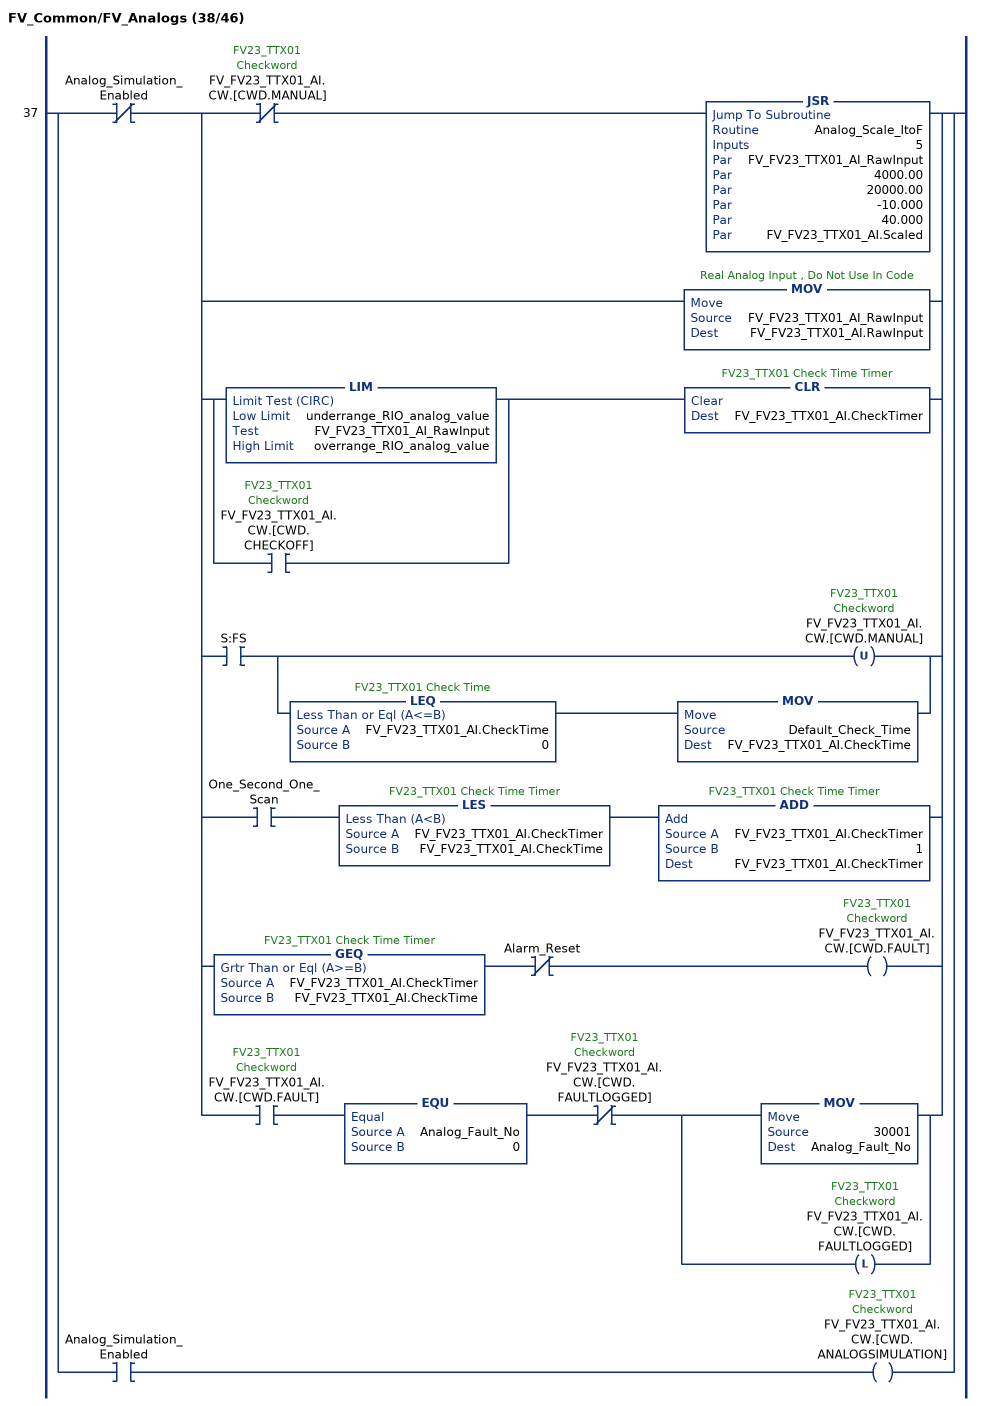
   37: [XIO(Analog_Simulation_Enabled) [XIO(FV_FV23_TTX01_AI.CW.[CWD.MANUAL]) JSR(Analog_Scale_ItoF,5,FV_FV23_TTX01_AI_RawInput,4000.00,20000.00,-10.000,40.000,FV_FV23_TTX01_AI.Scaled) ,MOV(FV_FV23_TTX01_AI_RawInput,FV_FV23_TTX01_AI.RawInput) ,[LIM(underrange_RIO_analog_value,FV_FV23_TTX01_AI_RawInput,overrange_RIO_analog_value) ,XIC(FV_FV23_TTX01_AI.CW.[CWD.CHECKOFF]) ] CLR(FV_FV23_TTX01_AI.CheckTimer) ,XIC(S:FS) [OTU(FV_FV23_TTX01_AI.CW.[CWD.MANUAL]) ,LEQ(FV_FV23_TTX01_AI.CheckTime,0) MOV(Default_Check_Time,FV_FV23_TTX01_AI.CheckTime) ] ,XIC(One_Second_One_Scan) LES(FV_FV23_TTX01_AI.CheckTimer,FV_FV23_TTX01_AI.CheckTime) ADD(FV_FV23_TTX01_AI.CheckTimer,1,FV_FV23_TTX01_AI.CheckTimer) ,GEQ(FV_FV23_TTX01_AI.CheckTimer,FV_FV23_TTX01_AI.CheckTime) XIO(Alarm_Reset) OTE(FV_FV23_TTX01_AI.CW.[CWD.FAULT]) ,XIC(FV_FV23_TTX01_AI.CW.[CWD.FAULT]) EQU(Analog_Fault_No,0) XIO(FV_FV23_TTX01_AI.CW.[CWD.FAULTLOGGED]) [MOV(30001,Analog_Fault_No) ,OTL(FV_FV23_TTX01_AI.CW.[CWD.FAULTLOGGED]) ] ] ,XIC(Analog_Simulation_Enabled) OTE(FV_FV23_TTX01_AI.CW.[CWD.ANALOGSIMULATION]) ];
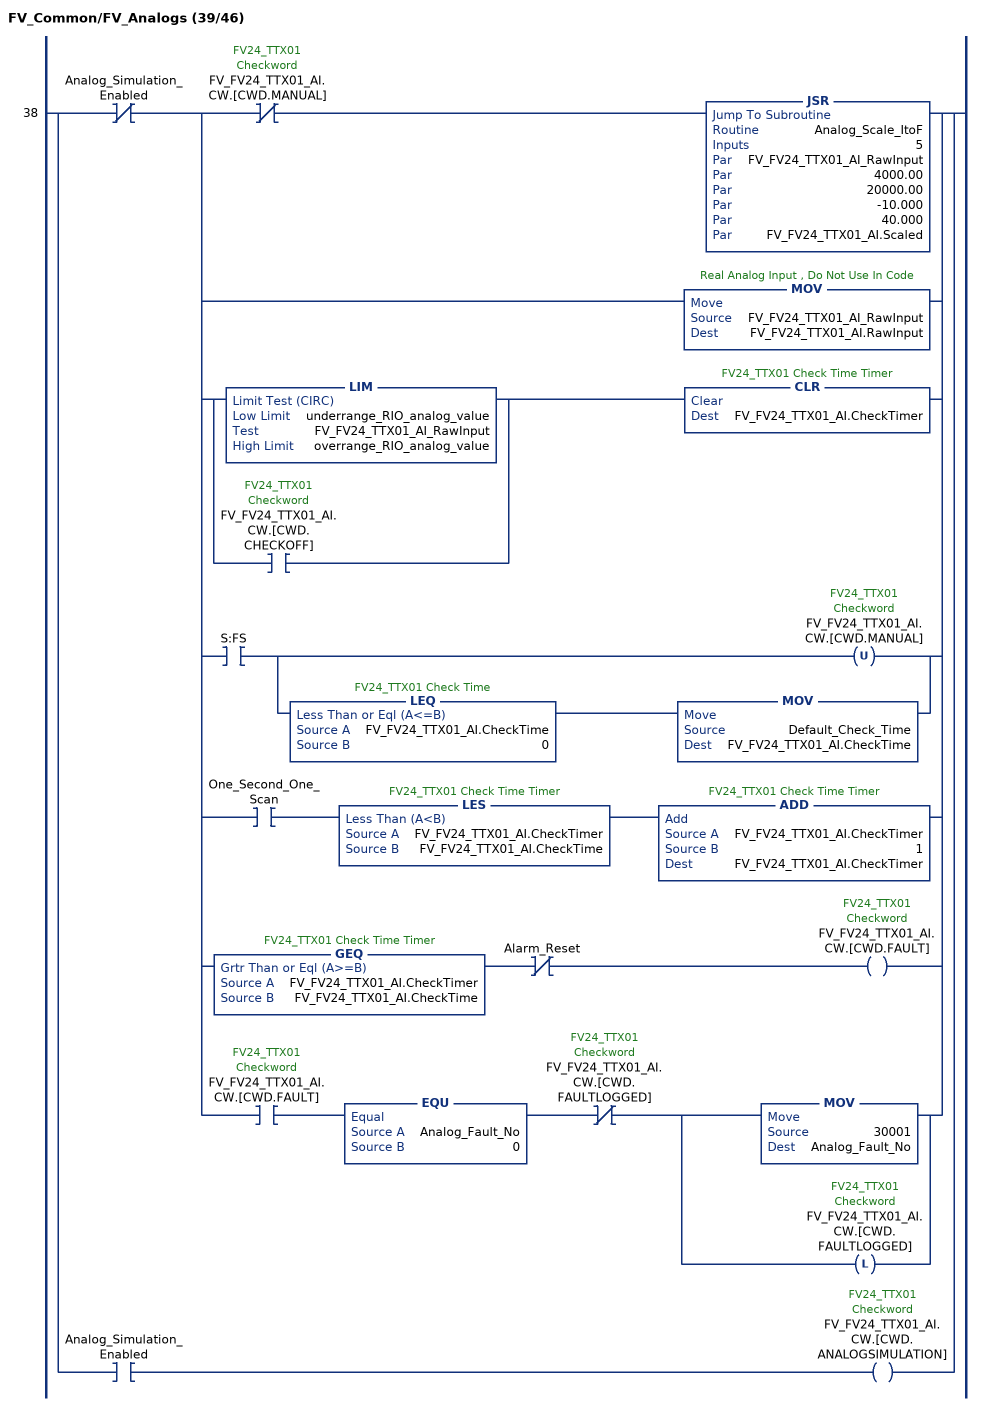
   38: [XIO(Analog_Simulation_Enabled) [XIO(FV_FV24_TTX01_AI.CW.[CWD.MANUAL]) JSR(Analog_Scale_ItoF,5,FV_FV24_TTX01_AI_RawInput,4000.00,20000.00,-10.000,40.000,FV_FV24_TTX01_AI.Scaled) ,MOV(FV_FV24_TTX01_AI_RawInput,FV_FV24_TTX01_AI.RawInput) ,[LIM(underrange_RIO_analog_value,FV_FV24_TTX01_AI_RawInput,overrange_RIO_analog_value) ,XIC(FV_FV24_TTX01_AI.CW.[CWD.CHECKOFF]) ] CLR(FV_FV24_TTX01_AI.CheckTimer) ,XIC(S:FS) [OTU(FV_FV24_TTX01_AI.CW.[CWD.MANUAL]) ,LEQ(FV_FV24_TTX01_AI.CheckTime,0) MOV(Default_Check_Time,FV_FV24_TTX01_AI.CheckTime) ] ,XIC(One_Second_One_Scan) LES(FV_FV24_TTX01_AI.CheckTimer,FV_FV24_TTX01_AI.CheckTime) ADD(FV_FV24_TTX01_AI.CheckTimer,1,FV_FV24_TTX01_AI.CheckTimer) ,GEQ(FV_FV24_TTX01_AI.CheckTimer,FV_FV24_TTX01_AI.CheckTime) XIO(Alarm_Reset) OTE(FV_FV24_TTX01_AI.CW.[CWD.FAULT]) ,XIC(FV_FV24_TTX01_AI.CW.[CWD.FAULT]) EQU(Analog_Fault_No,0) XIO(FV_FV24_TTX01_AI.CW.[CWD.FAULTLOGGED]) [MOV(30001,Analog_Fault_No) ,OTL(FV_FV24_TTX01_AI.CW.[CWD.FAULTLOGGED]) ] ] ,XIC(Analog_Simulation_Enabled) OTE(FV_FV24_TTX01_AI.CW.[CWD.ANALOGSIMULATION]) ];
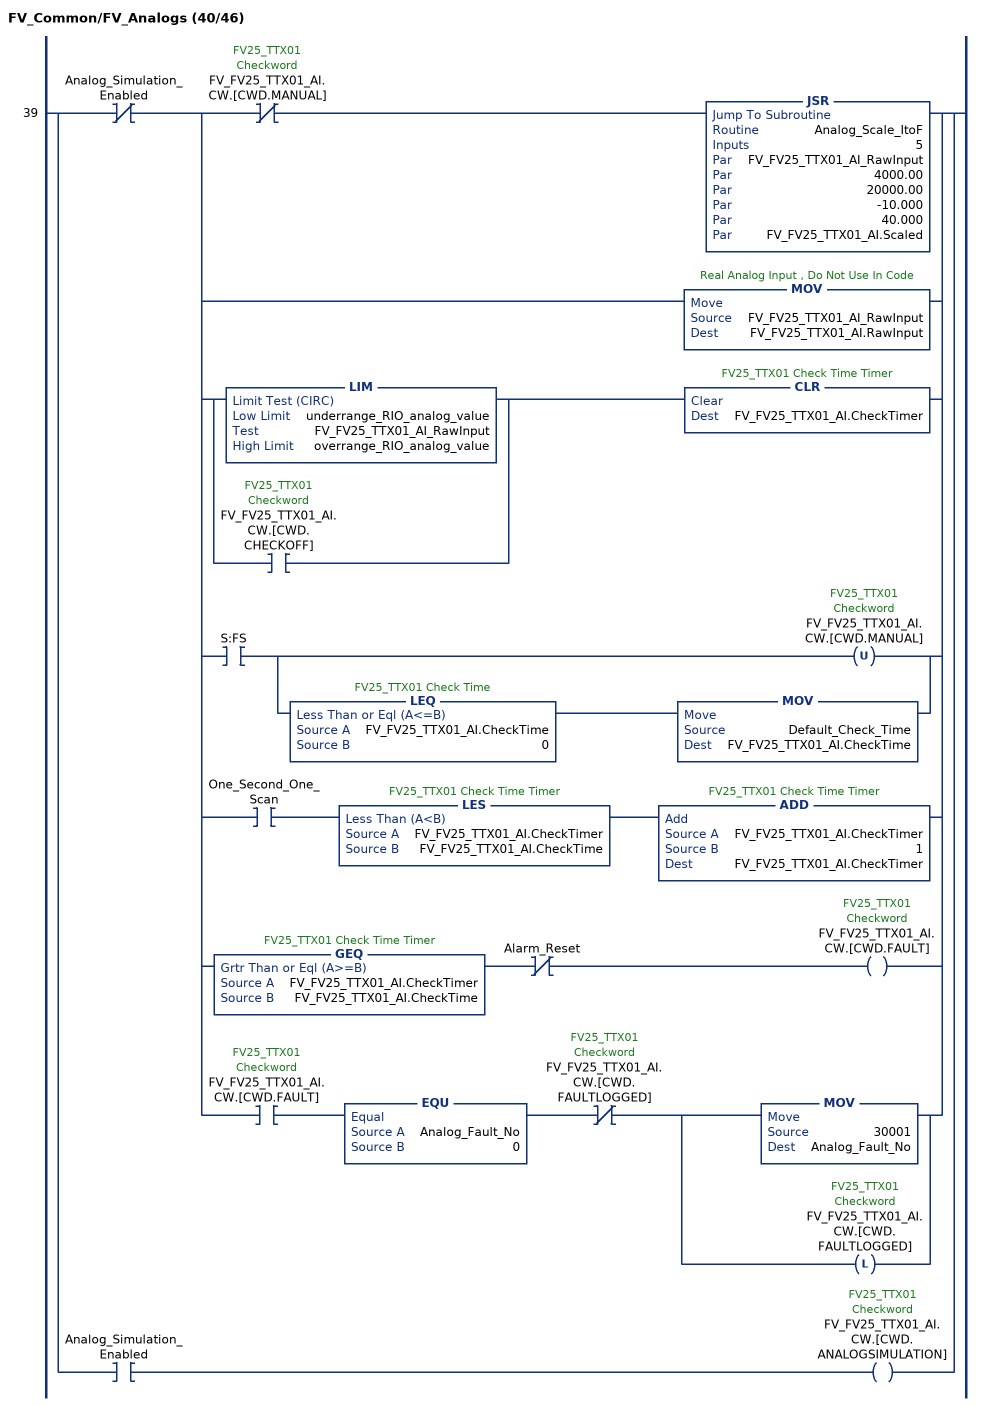
   39: [XIO(Analog_Simulation_Enabled) [XIO(FV_FV25_TTX01_AI.CW.[CWD.MANUAL]) JSR(Analog_Scale_ItoF,5,FV_FV25_TTX01_AI_RawInput,4000.00,20000.00,-10.000,40.000,FV_FV25_TTX01_AI.Scaled) ,MOV(FV_FV25_TTX01_AI_RawInput,FV_FV25_TTX01_AI.RawInput) ,[LIM(underrange_RIO_analog_value,FV_FV25_TTX01_AI_RawInput,overrange_RIO_analog_value) ,XIC(FV_FV25_TTX01_AI.CW.[CWD.CHECKOFF]) ] CLR(FV_FV25_TTX01_AI.CheckTimer) ,XIC(S:FS) [OTU(FV_FV25_TTX01_AI.CW.[CWD.MANUAL]) ,LEQ(FV_FV25_TTX01_AI.CheckTime,0) MOV(Default_Check_Time,FV_FV25_TTX01_AI.CheckTime) ] ,XIC(One_Second_One_Scan) LES(FV_FV25_TTX01_AI.CheckTimer,FV_FV25_TTX01_AI.CheckTime) ADD(FV_FV25_TTX01_AI.CheckTimer,1,FV_FV25_TTX01_AI.CheckTimer) ,GEQ(FV_FV25_TTX01_AI.CheckTimer,FV_FV25_TTX01_AI.CheckTime) XIO(Alarm_Reset) OTE(FV_FV25_TTX01_AI.CW.[CWD.FAULT]) ,XIC(FV_FV25_TTX01_AI.CW.[CWD.FAULT]) EQU(Analog_Fault_No,0) XIO(FV_FV25_TTX01_AI.CW.[CWD.FAULTLOGGED]) [MOV(30001,Analog_Fault_No) ,OTL(FV_FV25_TTX01_AI.CW.[CWD.FAULTLOGGED]) ] ] ,XIC(Analog_Simulation_Enabled) OTE(FV_FV25_TTX01_AI.CW.[CWD.ANALOGSIMULATION]) ];
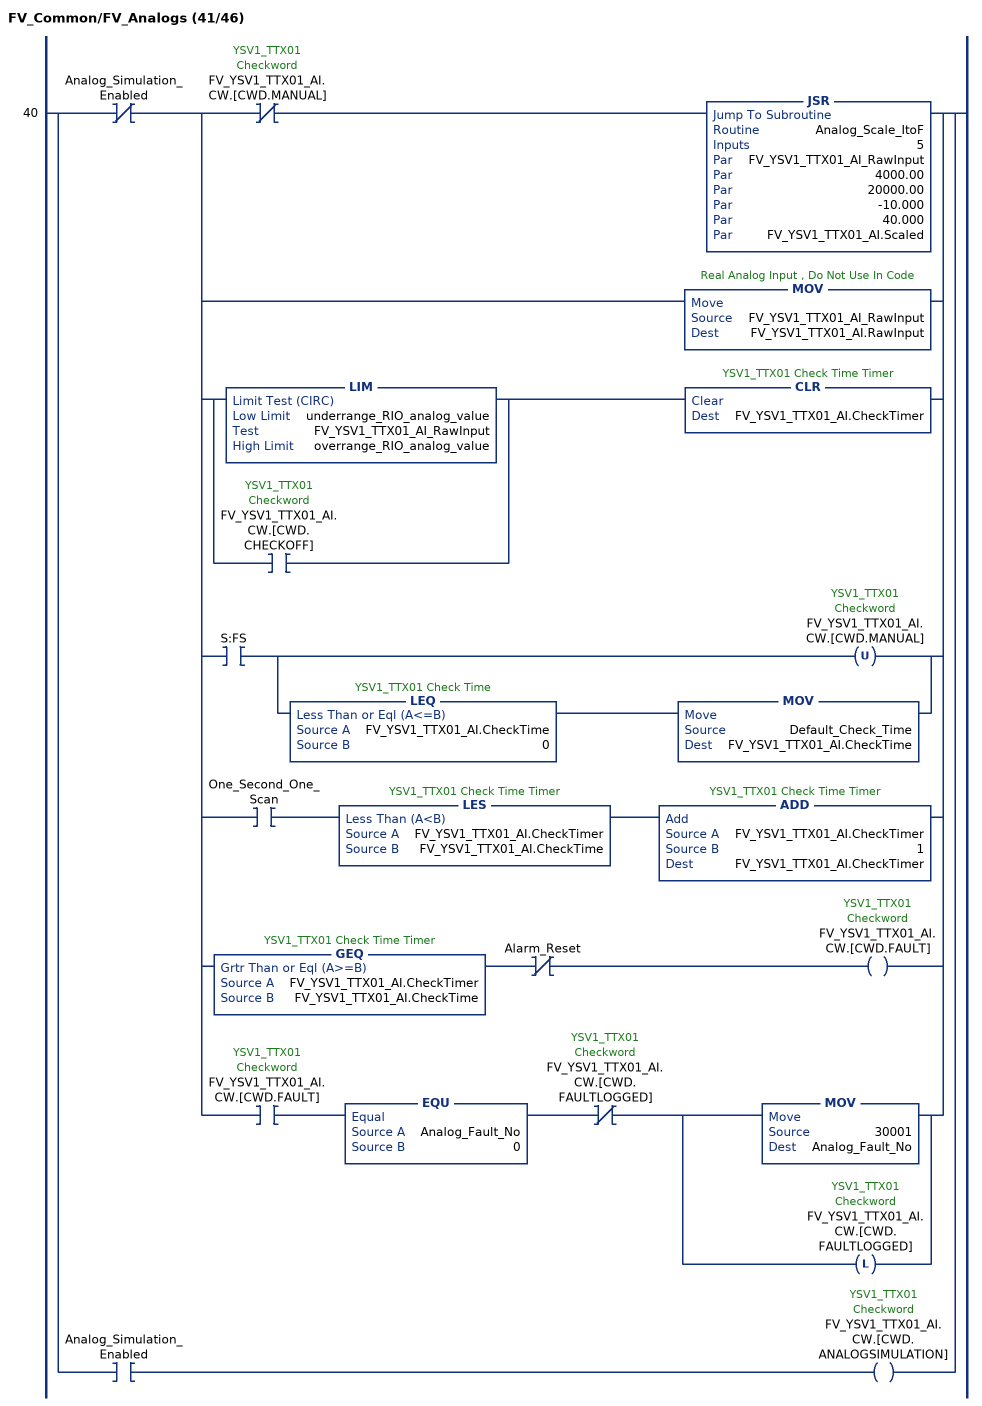
   40: [XIO(Analog_Simulation_Enabled) [XIO(FV_YSV1_TTX01_AI.CW.[CWD.MANUAL]) JSR(Analog_Scale_ItoF,5,FV_YSV1_TTX01_AI_RawInput,4000.00,20000.00,-10.000,40.000,FV_YSV1_TTX01_AI.Scaled) ,MOV(FV_YSV1_TTX01_AI_RawInput,FV_YSV1_TTX01_AI.RawInput) ,[LIM(underrange_RIO_analog_value,FV_YSV1_TTX01_AI_RawInput,overrange_RIO_analog_value) ,XIC(FV_YSV1_TTX01_AI.CW.[CWD.CHECKOFF]) ] CLR(FV_YSV1_TTX01_AI.CheckTimer) ,XIC(S:FS) [OTU(FV_YSV1_TTX01_AI.CW.[CWD.MANUAL]) ,LEQ(FV_YSV1_TTX01_AI.CheckTime,0) MOV(Default_Check_Time,FV_YSV1_TTX01_AI.CheckTime) ] ,XIC(One_Second_One_Scan) LES(FV_YSV1_TTX01_AI.CheckTimer,FV_YSV1_TTX01_AI.CheckTime) ADD(FV_YSV1_TTX01_AI.CheckTimer,1,FV_YSV1_TTX01_AI.CheckTimer) ,GEQ(FV_YSV1_TTX01_AI.CheckTimer,FV_YSV1_TTX01_AI.CheckTime) XIO(Alarm_Reset) OTE(FV_YSV1_TTX01_AI.CW.[CWD.FAULT]) ,XIC(FV_YSV1_TTX01_AI.CW.[CWD.FAULT]) EQU(Analog_Fault_No,0) XIO(FV_YSV1_TTX01_AI.CW.[CWD.FAULTLOGGED]) [MOV(30001,Analog_Fault_No) ,OTL(FV_YSV1_TTX01_AI.CW.[CWD.FAULTLOGGED]) ] ] ,XIC(Analog_Simulation_Enabled) OTE(FV_YSV1_TTX01_AI.CW.[CWD.ANALOGSIMULATION]) ];
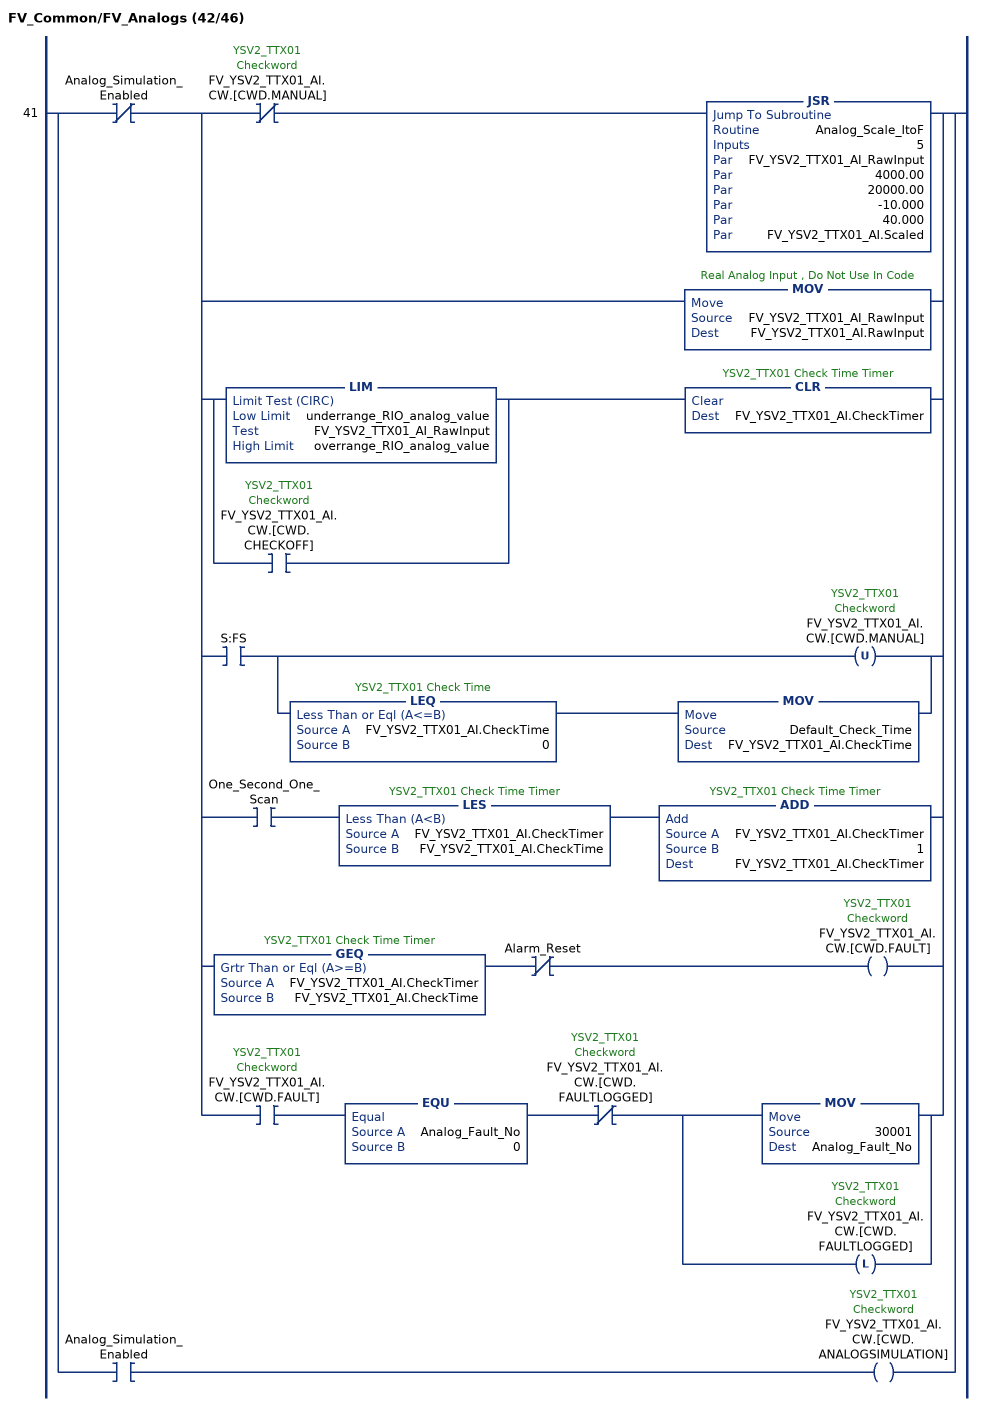
   41: [XIO(Analog_Simulation_Enabled) [XIO(FV_YSV2_TTX01_AI.CW.[CWD.MANUAL]) JSR(Analog_Scale_ItoF,5,FV_YSV2_TTX01_AI_RawInput,4000.00,20000.00,-10.000,40.000,FV_YSV2_TTX01_AI.Scaled) ,MOV(FV_YSV2_TTX01_AI_RawInput,FV_YSV2_TTX01_AI.RawInput) ,[LIM(underrange_RIO_analog_value,FV_YSV2_TTX01_AI_RawInput,overrange_RIO_analog_value) ,XIC(FV_YSV2_TTX01_AI.CW.[CWD.CHECKOFF]) ] CLR(FV_YSV2_TTX01_AI.CheckTimer) ,XIC(S:FS) [OTU(FV_YSV2_TTX01_AI.CW.[CWD.MANUAL]) ,LEQ(FV_YSV2_TTX01_AI.CheckTime,0) MOV(Default_Check_Time,FV_YSV2_TTX01_AI.CheckTime) ] ,XIC(One_Second_One_Scan) LES(FV_YSV2_TTX01_AI.CheckTimer,FV_YSV2_TTX01_AI.CheckTime) ADD(FV_YSV2_TTX01_AI.CheckTimer,1,FV_YSV2_TTX01_AI.CheckTimer) ,GEQ(FV_YSV2_TTX01_AI.CheckTimer,FV_YSV2_TTX01_AI.CheckTime) XIO(Alarm_Reset) OTE(FV_YSV2_TTX01_AI.CW.[CWD.FAULT]) ,XIC(FV_YSV2_TTX01_AI.CW.[CWD.FAULT]) EQU(Analog_Fault_No,0) XIO(FV_YSV2_TTX01_AI.CW.[CWD.FAULTLOGGED]) [MOV(30001,Analog_Fault_No) ,OTL(FV_YSV2_TTX01_AI.CW.[CWD.FAULTLOGGED]) ] ] ,XIC(Analog_Simulation_Enabled) OTE(FV_YSV2_TTX01_AI.CW.[CWD.ANALOGSIMULATION]) ];
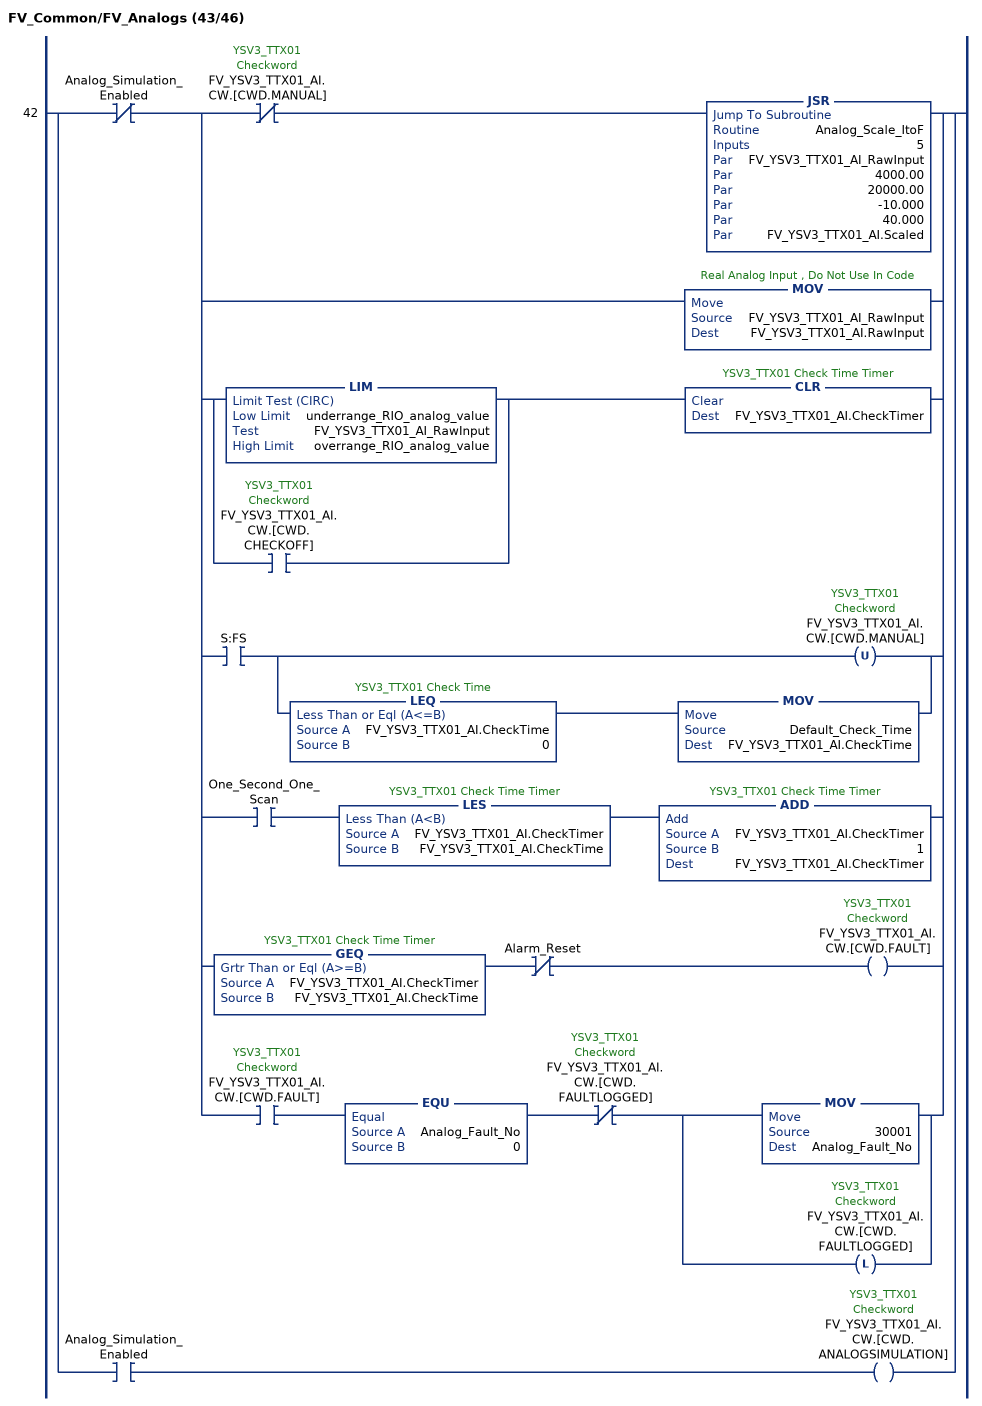
   42: [XIO(Analog_Simulation_Enabled) [XIO(FV_YSV3_TTX01_AI.CW.[CWD.MANUAL]) JSR(Analog_Scale_ItoF,5,FV_YSV3_TTX01_AI_RawInput,4000.00,20000.00,-10.000,40.000,FV_YSV3_TTX01_AI.Scaled) ,MOV(FV_YSV3_TTX01_AI_RawInput,FV_YSV3_TTX01_AI.RawInput) ,[LIM(underrange_RIO_analog_value,FV_YSV3_TTX01_AI_RawInput,overrange_RIO_analog_value) ,XIC(FV_YSV3_TTX01_AI.CW.[CWD.CHECKOFF]) ] CLR(FV_YSV3_TTX01_AI.CheckTimer) ,XIC(S:FS) [OTU(FV_YSV3_TTX01_AI.CW.[CWD.MANUAL]) ,LEQ(FV_YSV3_TTX01_AI.CheckTime,0) MOV(Default_Check_Time,FV_YSV3_TTX01_AI.CheckTime) ] ,XIC(One_Second_One_Scan) LES(FV_YSV3_TTX01_AI.CheckTimer,FV_YSV3_TTX01_AI.CheckTime) ADD(FV_YSV3_TTX01_AI.CheckTimer,1,FV_YSV3_TTX01_AI.CheckTimer) ,GEQ(FV_YSV3_TTX01_AI.CheckTimer,FV_YSV3_TTX01_AI.CheckTime) XIO(Alarm_Reset) OTE(FV_YSV3_TTX01_AI.CW.[CWD.FAULT]) ,XIC(FV_YSV3_TTX01_AI.CW.[CWD.FAULT]) EQU(Analog_Fault_No,0) XIO(FV_YSV3_TTX01_AI.CW.[CWD.FAULTLOGGED]) [MOV(30001,Analog_Fault_No) ,OTL(FV_YSV3_TTX01_AI.CW.[CWD.FAULTLOGGED]) ] ] ,XIC(Analog_Simulation_Enabled) OTE(FV_YSV3_TTX01_AI.CW.[CWD.ANALOGSIMULATION]) ];
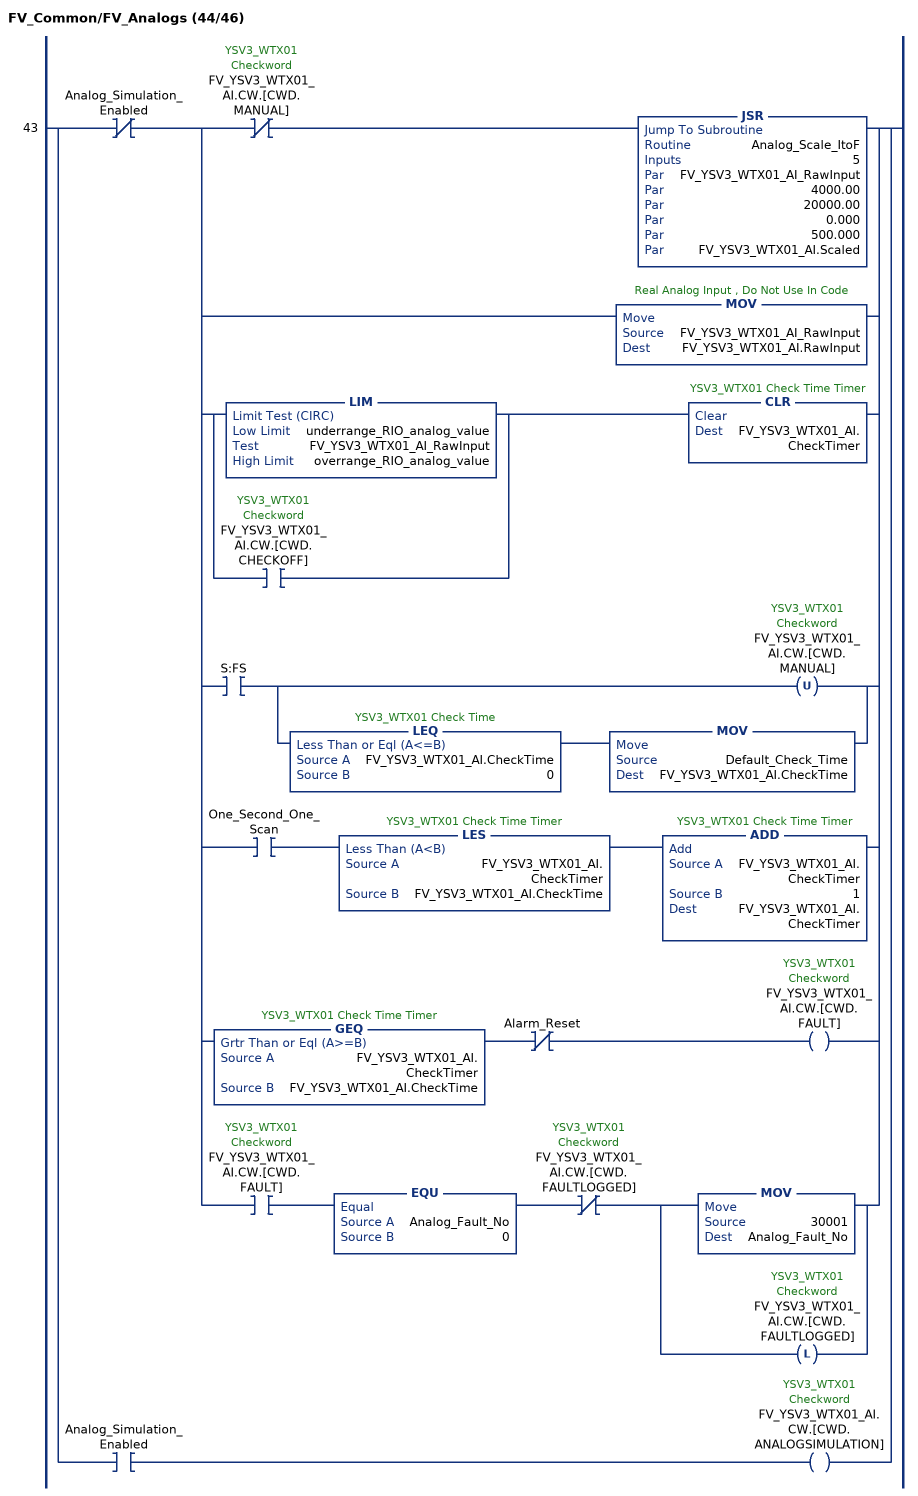
   43: [XIO(Analog_Simulation_Enabled) [XIO(FV_YSV3_WTX01_AI.CW.[CWD.MANUAL]) JSR(Analog_Scale_ItoF,5,FV_YSV3_WTX01_AI_RawInput,4000.00,20000.00,0.000,500.000,FV_YSV3_WTX01_AI.Scaled) ,MOV(FV_YSV3_WTX01_AI_RawInput,FV_YSV3_WTX01_AI.RawInput) ,[LIM(underrange_RIO_analog_value,FV_YSV3_WTX01_AI_RawInput,overrange_RIO_analog_value) ,XIC(FV_YSV3_WTX01_AI.CW.[CWD.CHECKOFF]) ] CLR(FV_YSV3_WTX01_AI.CheckTimer) ,XIC(S:FS) [OTU(FV_YSV3_WTX01_AI.CW.[CWD.MANUAL]) ,LEQ(FV_YSV3_WTX01_AI.CheckTime,0) MOV(Default_Check_Time,FV_YSV3_WTX01_AI.CheckTime) ] ,XIC(One_Second_One_Scan) LES(FV_YSV3_WTX01_AI.CheckTimer,FV_YSV3_WTX01_AI.CheckTime) ADD(FV_YSV3_WTX01_AI.CheckTimer,1,FV_YSV3_WTX01_AI.CheckTimer) ,GEQ(FV_YSV3_WTX01_AI.CheckTimer,FV_YSV3_WTX01_AI.CheckTime) XIO(Alarm_Reset) OTE(FV_YSV3_WTX01_AI.CW.[CWD.FAULT]) ,XIC(FV_YSV3_WTX01_AI.CW.[CWD.FAULT]) EQU(Analog_Fault_No,0) XIO(FV_YSV3_WTX01_AI.CW.[CWD.FAULTLOGGED]) [MOV(30001,Analog_Fault_No) ,OTL(FV_YSV3_WTX01_AI.CW.[CWD.FAULTLOGGED]) ] ] ,XIC(Analog_Simulation_Enabled) OTE(FV_YSV3_WTX01_AI.CW.[CWD.ANALOGSIMULATION]) ];
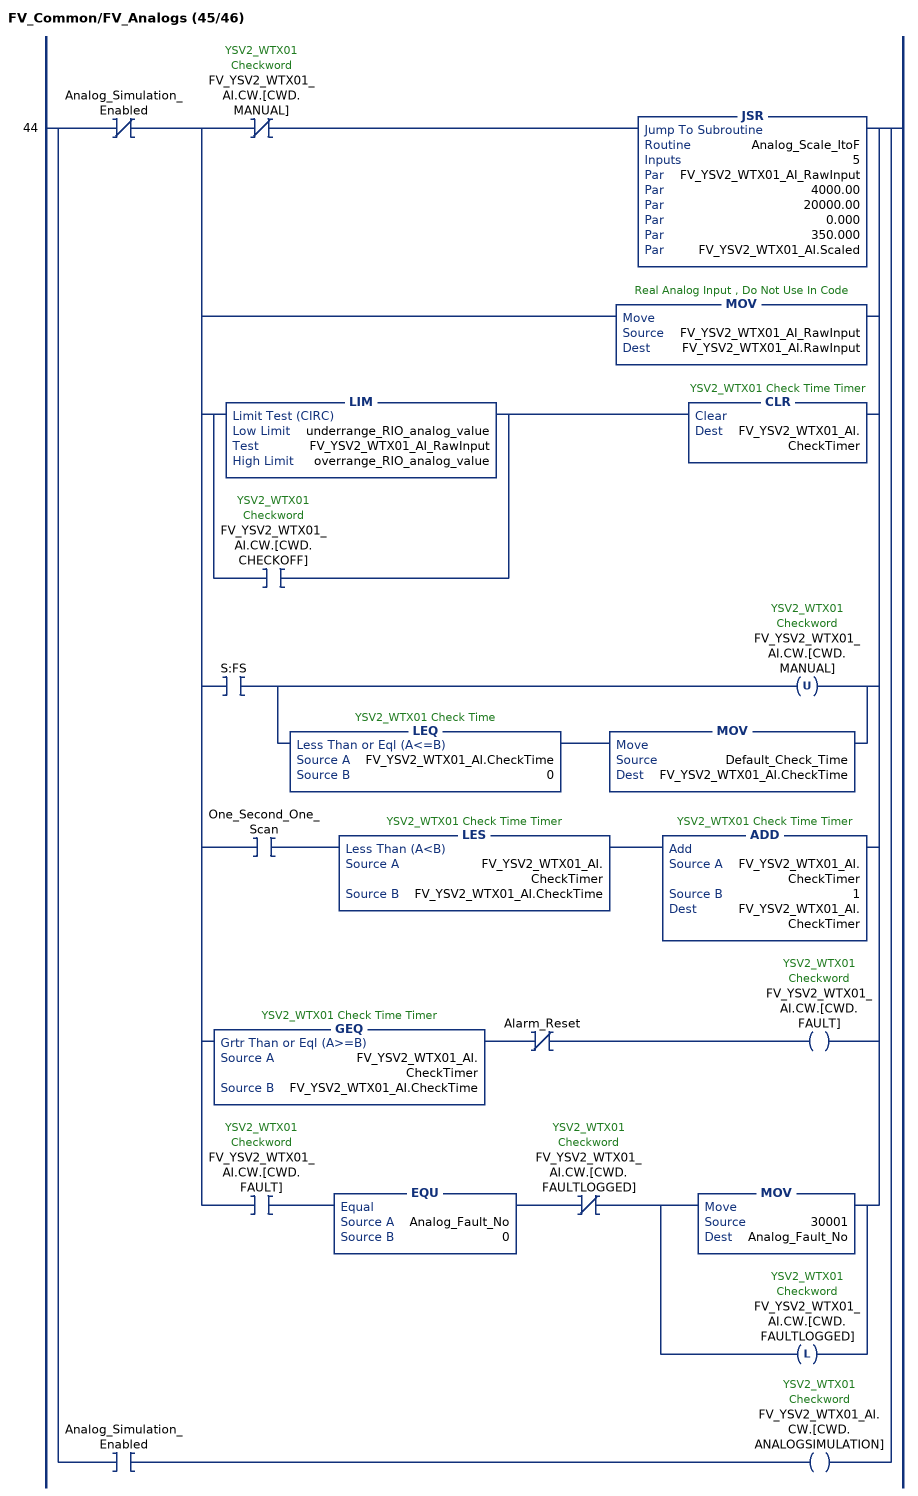
   44: [XIO(Analog_Simulation_Enabled) [XIO(FV_YSV2_WTX01_AI.CW.[CWD.MANUAL]) JSR(Analog_Scale_ItoF,5,FV_YSV2_WTX01_AI_RawInput,4000.00,20000.00,0.000,350.000,FV_YSV2_WTX01_AI.Scaled) ,MOV(FV_YSV2_WTX01_AI_RawInput,FV_YSV2_WTX01_AI.RawInput) ,[LIM(underrange_RIO_analog_value,FV_YSV2_WTX01_AI_RawInput,overrange_RIO_analog_value) ,XIC(FV_YSV2_WTX01_AI.CW.[CWD.CHECKOFF]) ] CLR(FV_YSV2_WTX01_AI.CheckTimer) ,XIC(S:FS) [OTU(FV_YSV2_WTX01_AI.CW.[CWD.MANUAL]) ,LEQ(FV_YSV2_WTX01_AI.CheckTime,0) MOV(Default_Check_Time,FV_YSV2_WTX01_AI.CheckTime) ] ,XIC(One_Second_One_Scan) LES(FV_YSV2_WTX01_AI.CheckTimer,FV_YSV2_WTX01_AI.CheckTime) ADD(FV_YSV2_WTX01_AI.CheckTimer,1,FV_YSV2_WTX01_AI.CheckTimer) ,GEQ(FV_YSV2_WTX01_AI.CheckTimer,FV_YSV2_WTX01_AI.CheckTime) XIO(Alarm_Reset) OTE(FV_YSV2_WTX01_AI.CW.[CWD.FAULT]) ,XIC(FV_YSV2_WTX01_AI.CW.[CWD.FAULT]) EQU(Analog_Fault_No,0) XIO(FV_YSV2_WTX01_AI.CW.[CWD.FAULTLOGGED]) [MOV(30001,Analog_Fault_No) ,OTL(FV_YSV2_WTX01_AI.CW.[CWD.FAULTLOGGED]) ] ] ,XIC(Analog_Simulation_Enabled) OTE(FV_YSV2_WTX01_AI.CW.[CWD.ANALOGSIMULATION]) ];
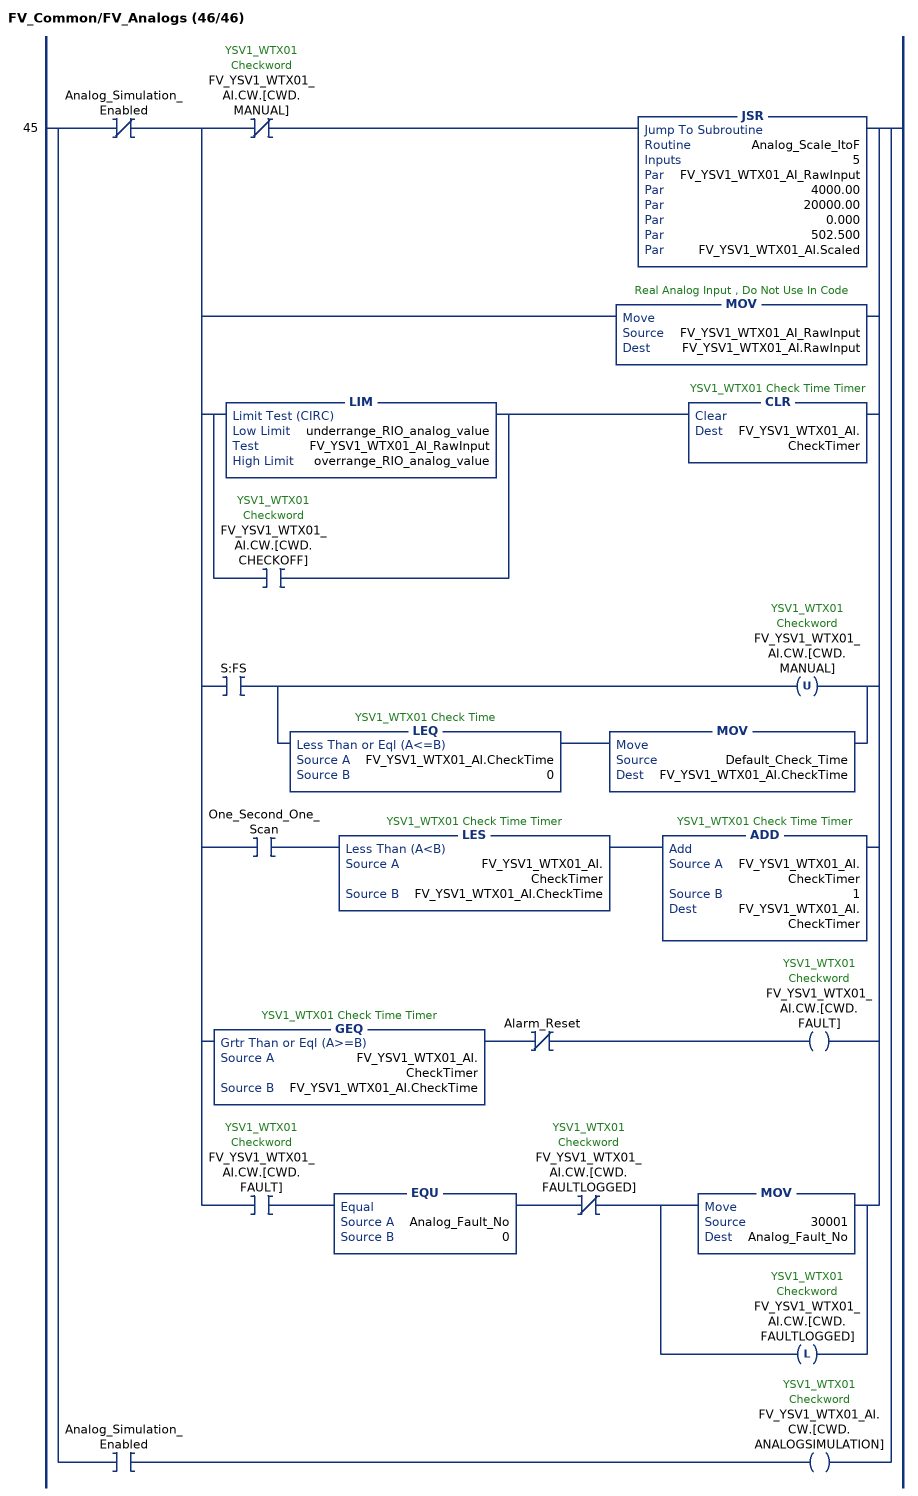
   45: [XIO(Analog_Simulation_Enabled) [XIO(FV_YSV1_WTX01_AI.CW.[CWD.MANUAL]) JSR(Analog_Scale_ItoF,5,FV_YSV1_WTX01_AI_RawInput,4000.00,20000.00,0.000,502.500,FV_YSV1_WTX01_AI.Scaled) ,MOV(FV_YSV1_WTX01_AI_RawInput,FV_YSV1_WTX01_AI.RawInput) ,[LIM(underrange_RIO_analog_value,FV_YSV1_WTX01_AI_RawInput,overrange_RIO_analog_value) ,XIC(FV_YSV1_WTX01_AI.CW.[CWD.CHECKOFF]) ] CLR(FV_YSV1_WTX01_AI.CheckTimer) ,XIC(S:FS) [OTU(FV_YSV1_WTX01_AI.CW.[CWD.MANUAL]) ,LEQ(FV_YSV1_WTX01_AI.CheckTime,0) MOV(Default_Check_Time,FV_YSV1_WTX01_AI.CheckTime) ] ,XIC(One_Second_One_Scan) LES(FV_YSV1_WTX01_AI.CheckTimer,FV_YSV1_WTX01_AI.CheckTime) ADD(FV_YSV1_WTX01_AI.CheckTimer,1,FV_YSV1_WTX01_AI.CheckTimer) ,GEQ(FV_YSV1_WTX01_AI.CheckTimer,FV_YSV1_WTX01_AI.CheckTime) XIO(Alarm_Reset) OTE(FV_YSV1_WTX01_AI.CW.[CWD.FAULT]) ,XIC(FV_YSV1_WTX01_AI.CW.[CWD.FAULT]) EQU(Analog_Fault_No,0) XIO(FV_YSV1_WTX01_AI.CW.[CWD.FAULTLOGGED]) [MOV(30001,Analog_Fault_No) ,OTL(FV_YSV1_WTX01_AI.CW.[CWD.FAULTLOGGED]) ] ] ,XIC(Analog_Simulation_Enabled) OTE(FV_YSV1_WTX01_AI.CW.[CWD.ANALOGSIMULATION]) ];
END_ROUTINE
